
   (* parse the format string *)
   #tDT_TO_STRF := #FMT;
   #pos := FIND(IN1:=#tDT_TO_STRF, IN2:='#');
   WHILE #pos > 0 DO
       (* retrieve format identifier *)
       #f := BYTE_TO_INT("CODE"(STR:=#tDT_TO_STRF, POS:=#pos + 1));
       (* generate the return string according to the format character *)
       #fs := '';
       CASE #f OF
           65 : (* letter A retunrs the year in 4 digits *)
               #fs := DELETE(IN:=S_CONV("YEAR_OF_DATE"(#dx)),L:=1,P:=1);
           66 : (* letter B returns the year in exactly 2 digits *)
               #fs := RIGHT(IN:=DELETE(IN:=S_CONV("YEAR_OF_DATE"(#dx)),L:=1,P:=1),L:=2);
           67 : (* letter C returns the month with 1 or 2 digits *)
               #fs := DELETE(IN:=S_CONV("MONTH_OF_DATE"(#dx)),L:=1,P:=1);
           68 : (* letter D returns the month with exactly 2 digits *)
               #fs := DELETE(IN:=S_CONV("MONTH_OF_DATE"(#dx)),L:=1,P:=1);
               IF LEN(#fs) < 2 THEN #fs := CONCAT(IN1:='0',IN2:=#fs); END_IF;
           69 : (* letter E returns the month with 3 characters *)
               #fs := "MONTH_TO_STRING"(MTH:="MONTH_OF_DATE"(#dx), LANG:=#ly, LX:=3);
           70 : (* letter F returns the month with all characters *)
               #fs := "MONTH_TO_STRING"(MTH:="MONTH_OF_DATE"(#dx), LANG:=#ly, LX:=0);
           71 : (* letter G returns the day with up to 2 digits *)
               #fs := DELETE(IN:=S_CONV("DAY_OF_MONTH"(#dx)),L:=1,P:=1);
           72 : (* letter H returns the day of the month with exactly 2 digits *)
               #fs := DELETE(IN:=S_CONV("DAY_OF_MONTH"(#dx)),L:=1,P:=1);
               IF LEN(#fs) < 2 THEN #fs := CONCAT(IN1:="FILL_FC235", IN2:=#fs); END_IF;
           73 : (* letter I returns the weekday as the number 1..7 1 = monday *)
               #fs := DELETE(IN:=S_CONV("DAY_OF_WEEK"(#dx)),L:=1,P:=1);
           74 : (* letter J returns the weekday in 2 character writing *)
               #fs := "WEEKDAY_TO_STRING"(WDAY:="DAY_OF_WEEK"(#dx), LANG:=#ly, LX:=2);
           75 : (* letter K returns the weekday with all characters *)
               #fs := "WEEKDAY_TO_STRING"(WDAY:="DAY_OF_WEEK"(#dx), LANG:=#ly, LX:=0);
           76 : (* letter L returns AM or PM for the given DateTime *)
               IF #td >= TOD#12:00:00 THEN #fs := 'PM'; ELSE #fs := 'AM'; END_IF;
           77 : (* letter M returns the hour in 1 or 2 digit form 0..24h *)
               #fs := DELETE(IN:=S_CONV("HOUR"(#td)),L:=1,P:=1);
           78 : (* letter N returns the hour in exactly 2 digit form 0..24h *)
               #fs := DELETE(IN:=S_CONV("HOUR"(#td)),L:=1,P:=1);
               IF LEN(#fs) < 2 THEN #fs := CONCAT(IN1:="FILL_FC235", IN2:=#fs); END_IF;
           79 : (* letter O returns the hour in 1 or 2 digit form 0..12h *)
               #tmp := "HOUR"(#td) MOD 12;
               IF #tmp = 0 THEN #tmp := 12; END_IF;
               #fs := DELETE(IN:=S_CONV(#tmp),L:=1,P:=1);
           80 : (* letter P returns the hour in exactly 2 digit form 0..12h *)
               #tmp := "HOUR"(#td) MOD 12;
               IF #tmp = 0 THEN #tmp := 12; END_IF;
               #fs := DELETE(IN:=S_CONV(#tmp),L:=1,P:=1);
               IF LEN(#fs) < 2 THEN #fs := CONCAT(IN1:="FILL_FC235", IN2:=#fs); END_IF;
           81 : (* letter Q returns the minute of the hour in 1 or two digit form *)
               #fs := DELETE(IN:=S_CONV("MINUTE"(#td)),L:=1,P:=1);
           82 : (* letter R returns the minute of the hour in exactly two digit form *)
               #fs := DELETE(IN:=S_CONV("MINUTE"(#td)),L:=1,P:=1);
               IF LEN(#fs) < 2 THEN #fs := CONCAT(IN1:="FILL_FC235", IN2:=#fs); END_IF;
           83 : (* letter S returns the second of the minute in 1 or two digit form *)
               #fs := DELETE(IN:=S_CONV(REAL_TO_INT("SECOND"(#td))),L:=1,P:=1);
           84 : (* letter T returns the second of the minute in exactly two digit form *)
               #fs := DELETE(IN:=S_CONV(REAL_TO_INT("SECOND"(#td))),L:=1,P:=1);
               IF LEN(#fs) < 2 THEN #fs := CONCAT(IN1:="FILL_FC235", IN2:=#fs); END_IF;
           85 : (* letter U returns the milliseconds in 1 to 3 digits *)
               #fs := DELETE(IN:=S_CONV(#MS),L:=1,P:=1);
           86 : (* letter V returns the milliseconds in exactly 3 digit form *)
               #fs := DELETE(IN:=S_CONV(#MS),L:=1,P:=1);
               #fs := CONCAT(IN1:='00',IN2:=#fs);
               #fs := RIGHT(IN:=#fs, L:=3);
           87 : (* letter W returns the day of the month with exactly 2 digits first digit is filled with blank if necessary *)
               #fs := DELETE(IN:=S_CONV("DAY_OF_MONTH"(#dx)),L:=1,P:=1);
               IF LEN(#fs) < 2 THEN #fs := CONCAT(IN1:="BLANK", IN2:=#fs); END_IF;
           88 : (* letter X returns the month with exactly 2 digits first digit is filled with blank if necessary *)
               #fs := DELETE(IN:=S_CONV("MONTH_OF_DATE"(#dx)),L:=1,P:=1);
               IF LEN(#fs) < 2 THEN #fs := CONCAT(IN1:="BLANK", IN2:=#fs); END_IF;
           END_CASE;
       #tDT_TO_STRF := REPLACE(IN1:=#tDT_TO_STRF, IN2:=#fs, L:=2, P:=#pos);
       #pos := FIND(IN1:=#tDT_TO_STRF, IN2:='#');
   END_WHILE;

   #DT_TO_STRF := #tDT_TO_STRF;

   (* revision history
   hm  7. oct. 2008    rev 1.0
       original version

   hm  19. oct. 2008   rev 1.1
       changed language setup constants
   *)
END_FUNCTION

FUNCTION "DWORD_TO_STRB" : String[254]   // FC236, SCL
TITLE = DWORD_TO_STRB
{ S7_Optimized_Access := 'FALSE' }
AUTHOR : hugo
FAMILY : STRINGS
NAME : DW2STRB
VERSION : 1.3
// DWORD_TO_STRINGB converts a DWORD to a String of Bits represented by '0' and '1' s.
// The lowest order bit will be on the right and the high order bit on the left.
   VAR_INPUT
      IN : DWord;
   END_VAR
   VAR_TEMP
      pt : Int;   // pt : POINTER TO BYTE;
      i : Int;
      str : String[32];
      _str AT str : Struct
         length : Byte;
         act_length : Byte;
         str : Array[1..32] of Byte;
      END_STRUCT;
      tIN : DWord;
      _IN AT tIN : Array[0..31] of Bool;
   END_VAR
BEGIN


   #str := #DWORD_TO_STRB;
   #tIN := #IN;

   (* pointer für die ausgabe ermitteln *)
   #pt := 1;    //ADR(DWORD_TO_STRB);
   (* die 8 ausgabecharacter ermitteln und schreiben *)
   FOR #i := 1 TO 32 DO
       #_str.str[#pt] := INT_TO_BYTE(BYTE_TO_INT(BOOL_TO_BYTE(#_IN[7])) + 48);
       #tIN := SHL(IN:=#tIN,N:=1);
       #pt := #pt + 1;
   END_FOR;

   (* der ausgabestring muss nochg mit 32 abgeschlossen werden *)
   #_str.act_length := 32;
   #DWORD_TO_STRB := #str;

   (* revision history
   hm      9.6.2007    rev 1.0     
       original version

   hm      15.dec 2007 rev 1.1
       changed code for better performance

   hm  29. mar. 2008   rev 1.2
       changed STRING to STRING(32)

   hm  20. jun. 2008   rev 1.3
       performance improvement

   *)
END_FUNCTION

FUNCTION "DWORD_TO_STRF" : String[254]   // FC237, SCL
TITLE = DWORD_TO_STRF
{ S7_Optimized_Access := 'FALSE' }
AUTHOR : hugo
FAMILY : STRINGS
NAME : DW2STRF
VERSION : 1.1
// dword_to_strF converts a DWORD, BYTE or Word to a fixed length String.
// the string will be filled with leading zeroes to achieve the fixed length, or if too long, the lowest digits will be used.
// the maximum allowed length is 20 mdigits.
//  
// for example:    dword_to_strf(123,4) = '0123' 
//                 dword_to_strf(123,2) = '23'
// 
// uses: CONCAT [FC2]
//       DI_STRNG [FC5]
//       MID [FC26]
//       LEN [FC21]
   VAR_INPUT
      IN : DWord;
      N : Int;
   END_VAR
   VAR_TEMP
      L : Int;
      temp : String[10];
      temp2 : String[10];
   END_VAR
BEGIN


   (* convert dword to string first and cut to length N *)
   #temp := '0';
   #temp2 := '0';
   #temp := MID(IN:=S_CONV(DWORD_TO_DINT(#IN)), L:=#N, P:=2);
   #L := LEN(#temp);

   WHILE #L < #N DO
       #temp2 := CONCAT(IN1:='0',IN2:=#temp);
       #temp BLKMOV #temp2;
       #L := #L + 1;
   END_WHILE;
   #DWORD_TO_STRF := #temp;


   (* limit N to max 20 characters *)
   //tN := LIMIT(IN1:=0,IN2:=tN,IN3:=20);
   (* convert dword to string first and cut to length N *)
   //str := FIX(DWORD_TO_STRING(in),tN,48,1);

   (* revision history
   hm  26. jan.2007    rev 1.0     
       original version

   hm  29. mar. 2008   rev 1.1
       changed STRING to STRING(20)
       limit the output string to max 20 digits
   *)
END_FUNCTION

FUNCTION "DWORD_TO_STRH" : String[254]   // FC238, SCL
TITLE = DWORD_TO_STRH
{ S7_Optimized_Access := 'FALSE' }
AUTHOR : hugo
FAMILY : STRINGS
NAME : DW2STRH
VERSION : 1.3
// DWORD_TO_STRINGH converts a DWORD to a String of Hexadecimal represented by '0' .. '9' and 'A' .. 'F'.
// The lowest order Character will be on the right and the high order Character on the left.
   VAR_INPUT
      IN : DWord;
   END_VAR
   VAR_TEMP
      i : Int;
      temp : Byte;
      pt : Int;   // pt : POINTER TO BYTE;
      str : String[8];
      _str AT str : Struct
         length : Byte;
         act_length : Byte;
         str : Array[1..8] of Byte;
      END_STRUCT;
      tIN : DWord;
   END_VAR
BEGIN


   #str := #DWORD_TO_STRH;
   #tIN := #IN;

   (* read output adress to pointer *)
   #pt := 8;    //ADR(DWORD_TO_STRH) + 8;
   (* wirte the closing byte for the string *)
   //_str.str[pt]:= 0;

   (* write the 8 hex characters backwards *)
   FOR #i := 1 TO 8 DO;
       (* read the lowest order hex value *)
       #temp := DWORD_TO_BYTE(#tIN AND 16#0000000F);
       (* convert value to hex character *)
       IF BYTE_TO_INT(#temp) <= 9 THEN #temp := INT_TO_BYTE(BYTE_TO_INT(#temp) + 48); ELSE #temp := INT_TO_BYTE(BYTE_TO_INT(#temp) + 55); END_IF;
       (* write character to output string *)
       #_str.str[#pt] := #temp;
       (* shift in for nect hex character *)
       #tIN := SHR(IN:=#tIN,N:=4);
       (* decrement the pointer *)
       #pt := #pt - 1;
   END_FOR;

   #_str.act_length := 8;
   #DWORD_TO_STRH := #str;

   (* code beofre rev 1.2
   FOR i := 1 TO 8 DO
       X := DWORD_TO_BYTE(in AND 2#1111);
       IF X <= 9 THEN X := X + 48; ELSE X := X + 55; END_IF;
       Cx := CHR(X);
       temp := CONCAT(Cx, temp);
       in := SHR(in,4);
   END_FOR;
   DWORD_TO_STRH := temp;
   *)


   (* revision history
   hm  9. jun. 2007    rev 1.0     
       original version 

   hm  11. sep. 2007   rev 1.1
       changed coding for compatibility with twincat, concat cannot support a function as an argument.

   hm  15. dec. 2007    rev 1.2
       changed code for better performance

   hm  29. mar. 2008   rev 1.3
       changed STRING to STRING(8)

   *)
END_FUNCTION

FUNCTION "EXEC" : String[254]   // FC239, SCL
TITLE = EXEC
{ S7_Optimized_Access := 'FALSE' }
AUTHOR : hugo
FAMILY : STRINGS
NAME : EXEC
VERSION : 1.4
// exec executes a mathematical term and returns the result as a string
// the term can only be a simple term without brackets and only one operator
// allowed operastors are: (+, -, *, /, ^, sqrt, sin, cos, tan).
// 
// uses: SETUP [DB1]
//       TEMP [DB7]
//       EQ_STRNG [FC10]
//       R_STRNG [FC30]
//       STRNG_R [FC39]
//       CONCAT [FC2]
//       UPPERCASE [FC288]
//       TO_UPPER [FC284] 
//       TRIM [FC285]
//       FIND [FC11] 
//       REPLACE [FC31] 
//       FINDB_NONUM [FC246]
//       LEFT [FC20]
//       RIGHT [FC32]
//       LEN [FC21]
//       FINDB_NUM [FC247]
   VAR_INPUT
      str : String[254];
   END_VAR
   VAR_TEMP
      pos : Int;
      R1 : Real;
      R2 : Real;
      operator : String[10];
   END_VAR
BEGIN


   "TEMP".STR1 := #str;

   (* extract both numbers and operator *)
   "TEMP".STR2 := "UPPERCASE"("TRIM"("TEMP".STR1));

   #pos := "FINDB_NONUM"("TEMP".STR2);
   IF #pos > 1 THEN #R1 := S_CONV(LEFT(IN:="TEMP".STR2,L:=#pos-1)); END_IF;
   #R2 := S_CONV(RIGHT(IN:="TEMP".STR2,L:=LEN("TEMP".STR2)-#pos));
   "TEMP".STR2 := LEFT(IN:="TEMP".STR2,L:=#pos);
   #pos := "FINDB_NUM"("TEMP".STR2);
   #operator := RIGHT(IN:="TEMP".STR2,L:=LEN("TEMP".STR2) - #pos);
   IF #operator = '' AND LEN("TEMP".STR1) = 0 THEN
       #EXEC := '';
       RETURN;
   ELSIF #operator = '' THEN
       "TEMP".STR2 := "TEMP".STR1;
       RETURN;
   END_IF;
   IF #operator = '^' THEN
       "TEMP".STR2 := S_CONV((#R1**#R2));
   ELSIF #operator = 'SQRT' THEN
       "TEMP".STR2 := S_CONV(SQRT(#R2));
   ELSIF #operator = 'SIN' THEN
       "TEMP".STR2 := S_CONV(SIN(#R2));
   ELSIF #operator = 'COS' THEN
       "TEMP".STR2 := S_CONV(COS(#R2));
   ELSIF #operator = 'TAN' THEN
       "TEMP".STR2 := S_CONV(TAN(#R2));
   ELSIF #operator = '*' THEN
       "TEMP".STR2 := S_CONV(#R1 * #R2);
   ELSIF #operator = '/' THEN
       IF #R2 <> 0 THEN "TEMP".STR2 := S_CONV(#R1 / #R2); ELSE "TEMP".STR2 := 'ERROR'; END_IF;
   ELSIF #operator = '+' THEN
       "TEMP".STR2 := S_CONV(#R1 + #R2);
   ELSIF #operator = '-' THEN
       "TEMP".STR2 := S_CONV(#R1 - #R2);
   ELSE
       "TEMP".STR2 := 'ERROR';
   END_IF;

   IF "TEMP".STR2 = 'ERROR' THEN
       RETURN;
   (* some systems deliver integer instead of real *)
   ELSIF FIND(IN1:="TEMP".STR2,IN2:='.') = 0 THEN
       "TEMP".STR2 := CONCAT(IN1:="TEMP".STR2,IN2:='.0');
   (* some systems deliver n. instead of n.0 ! *)
   ELSIF RIGHT(IN:="TEMP".STR2,L:=1) = '.' THEN
       "TEMP".STR2 := CONCAT(IN1:="TEMP".STR2,IN2:='0');
   END_IF;

   #EXEC := "TEMP".STR2;

   (* revision history

   hm  6.feb 2007      rev 1.1
       cos has to be written in uppercase
       divide by 0 will return an error

   hm  5. mar. 2008    rev 1.2
       add a 0 to the string if a '.' is at the end of the string

   hm  20. mar. 2008   rev 1.3
       make sure the function always returns a real value in the form of x.y

   hm  29. mar. 2008   rev 1.4
       changed STRING to STRING(STRING_LENGTH)
   *)
END_FUNCTION

FUNCTION "FILL" : String[254]   // FC240, SCL
TITLE = FILL
{ S7_Optimized_Access := 'FALSE' }
AUTHOR : hugo
FAMILY : STRINGS
NAME : FILL
VERSION : 1.1
// the function fill creates a string at length L of characters C.
//  
// uses: CONSTANTS [DB6]
//       CONCAT [FC2]
//       CHR_TO_STRING [FC227]
   VAR_INPUT
      C : Byte;
      L : Int;
   END_VAR
   VAR_TEMP
      tFILL : String[254];
      tL : Word;
      _L AT tL : Array[0..15] of Bool;
      i : Int;
      sx : String[1];
   END_VAR
BEGIN


   #sx := "CHR_TO_STRING"(#C);
   (* limit L to maximum 80 characters the length of a standard string *)
   #tL := INT_TO_WORD(LIMIT(MN:=0,IN:=#L,MX:="CONSTANTS".STRING_LENGTH));
   (* create a string of characters to be connected to str *)
   FOR #i := 1 TO 8 DO
       #tFILL := CONCAT(IN1:=#tFILL,IN2:=#tFILL);
       IF #_L[15] THEN #tFILL := CONCAT(IN1:=#tFILL,IN2:=#sx); END_IF;
       #tL := SHL(IN:=#tL,N:=1);
   END_FOR;

   #FILL := #tFILL;


   (* revision histroy
   hm  29. mar. 2008   rev 1.0
       original release

   hm  17. dec. 2008   rev 1.1
       changed function chr to chr_to_string

   *)
END_FUNCTION

FUNCTION "FIND_CHAR" : Int   // FC241, SCL
TITLE = FIND_CHAR
{ S7_Optimized_Access := 'FALSE' }
AUTHOR : hugo
FAMILY : STRINGS
NAME : FCHAR
VERSION : 1.3
// find_char searches str and returns the starting position of the first character that is not a control character.
// control characters are the ascii character 00 .. 31.
// 
// uses: SETUP [DB1]
   VAR_INPUT
      str : String[254];
      _str AT str : Struct
         length : Byte;
         act_length : Byte;
         str : Array[1..254] of Byte;
      END_STRUCT;
      pos : Int;
   END_VAR
   VAR_TEMP
      i : Int;
      stop : Int;
      X : Byte;
   END_VAR
BEGIN


   #stop := BYTE_TO_INT(#_str.act_length);
   FOR #i := MAX(IN1:=#pos,IN2:=1) TO #stop DO
       #X := #_str.str[#i];
       IF BYTE_TO_INT(#X) > 31 AND (("SETUP".EXTENDED_ASCII AND BYTE_TO_INT(#X) <> 127) OR (NOT "SETUP".EXTENDED_ASCII AND BYTE_TO_INT(#X) < 127)) THEN
           #FIND_CHAR := #i;
           RETURN;
       END_IF;
   END_FOR;
   #FIND_CHAR := 0;


   (* revision history
   hm  29. feb 2008    rev 1.0
       original version

   hm  26. mar. 2008   rev 1.1
       char will now accept extended ascii

   hm  29. mar. 2008   rev 1.2
       changed STRING to STRING(STRING_LENGTH)

   hm  21. oct. 2008 rev 1.3
       changes setup constants
       optimized code
   *)
END_FUNCTION

FUNCTION "FIND_CTRL" : Int   // FC242, SCL
TITLE = FIND_CTRL
{ S7_Optimized_Access := 'FALSE' }
AUTHOR : hugo
FAMILY : STRINGS
NAME : FCTRL
VERSION : 1.2
// find_ctrl searches str and returns the starting position of a control character
// control characters are the ascii character 00 .. 31.
   VAR_INPUT
      str : String[254];
      _str AT str : Struct
         length : Byte;
         act_length : Byte;
         str : Array[1..254] of Byte;
      END_STRUCT;
      pos : Int;
   END_VAR
   VAR_TEMP
      i : Int;
      stop : Int;
      x : Byte;
   END_VAR
BEGIN


   #stop := BYTE_TO_INT(#_str.act_length);
   FOR #i := MAX(IN1:=#pos,IN2:=1) TO #stop DO;
       #x := #_str.str[#i];
       IF BYTE_TO_INT(#x) < 32 OR BYTE_TO_INT(#x) = 127 THEN
           #FIND_CTRL := #i;
           RETURN;
       END_IF;
   END_FOR;
   #FIND_CTRL := 0;


   (* revision history
   hm  29. feb 2008    rev 1.0
       original version

   hm  26. mar. 2008   rev 1.1
       character 127 is now recognized as control

   hm  29. mar. 2008   rev 1.2
       changed STRING to STRING(STRING_LENGTH)
   *)
END_FUNCTION

FUNCTION "FIND_NONUM" : Int   // FC243, SCL
TITLE = FIND_NONUM
{ S7_Optimized_Access := 'FALSE' }
AUTHOR : hugo
FAMILY : STRINGS
NAME : FINDNONR
VERSION : 1.3
// find_noNum searches str AND returns the first position which is NOT a number.
// a number is characterized by a letter "0..9" or "."
   VAR_INPUT
      str : String[254];
      _str AT str : Struct
         length : Byte;
         act_length : Byte;
         str : Array[1..254] of Byte;
      END_STRUCT;
      pos : Int;
   END_VAR
   VAR_TEMP
      i : Int;
      end : Int;
      X : Byte;
   END_VAR
BEGIN


   #end := BYTE_TO_INT(#_str.act_length);    //LEN(str);
   FOR #i := MAX(IN1:=#pos,IN2:=1) TO #end DO
       #X := #_str.str[#i];
       IF (BYTE_TO_INT(#X) < 48 AND BYTE_TO_INT(#X) <> 46) OR BYTE_TO_INT(#X) > 57 THEN
           #FIND_NONUM := #i;
           RETURN;
       END_IF;
   END_FOR;
   #FIND_NONUM := 0;


   (* revision history
   hm  6. oct. 2006    rev 1.0
       original version

   hm  29. feb 2008    rev 1.1
       added input pos to start search at position

   hm  29. mar. 2008   rev 1.2
       changed STRING to STRING(STRING_LENGTH)

   hm  21. oct. 2008   rev 1.3
       optimized code

   *)
END_FUNCTION

FUNCTION "FIND_NUM" : Int   // FC244, SCL
TITLE = FIND_NUM
{ S7_Optimized_Access := 'FALSE' }
AUTHOR : hugo
FAMILY : STRINGS
NAME : FINDNR
VERSION : 1.2
// find_Num searches str and returns the starting position of a number
// a number is characterized by a letter "0..9" or "."
   VAR_INPUT
      str : String[254];
      _str AT str : Struct
         length : Byte;
         act_length : Byte;
         str : Array[1..254] of Byte;
      END_STRUCT;
      pos : Int;
   END_VAR
   VAR_TEMP
      i : Int;
      stop : Int;
      X : Byte;
   END_VAR
BEGIN


   #stop := BYTE_TO_INT(#_str.act_length);   //LEN(str);
   FOR #i := MAX(IN1:=#pos,IN2:=1) TO #stop DO;
       #X := #_str.str[#i];
       IF (BYTE_TO_INT(#X) > 47 AND BYTE_TO_INT(#X) < 58) OR BYTE_TO_INT(#X) = 46 THEN
           #FIND_NUM := #i;
           RETURN;
       END_IF;
   END_FOR;
   #FIND_NUM := 0;


   (* revision history
   hm  6. oct. 2006    rev 1.0
       original version

   hm  29. feb 2008    rev 1.1
       added input pos to start search at position

   hm  29. mar. 2008   rev 1.2
       changed STRING to STRING(STRING_LENGTH)

   *)
END_FUNCTION

FUNCTION "FINDB" : Int   // FC245, SCL
TITLE = FINDB
{ S7_Optimized_Access := 'FALSE' }
AUTHOR : hugo
FAMILY : STRINGS
NAME : FINDB
VERSION : 1.3
// the function find searches an str1 for the presence of str2 and returns the first position of str1 of the last presence in instring.
// the function is similar to find except it searches from the right to left.
// a 0 is returned if the string is not found.
//  
// uses: EQ_STRNG [FC10]
//       MID [FC26]
   VAR_INPUT
      str1 : String[254];
      str2 : String[254];
   END_VAR
   VAR_TEMP
      tstr1 : String[254];
      _str1 AT tstr1 : Struct
         length : Byte;
         act_length : Byte;
         str : Array[1..254] of Byte;
      END_STRUCT;
      tstr2 : String[254];
      _str2 AT tstr2 : Struct
         length : Byte;
         act_length : Byte;
         str : Array[1..254] of Byte;
      END_STRUCT;
      pos : Int;
      length : Int;
   END_VAR
BEGIN


   #tstr1 := #str1;
   #tstr2 := #str2;

   #length := BYTE_TO_INT(#_str2.act_length);
   FOR #pos := BYTE_TO_INT(#_str1.act_length) - #length + 1 TO 1 BY -1 DO
       IF MID(IN:=#tstr1,L:=#length,P:=#pos) S_COMP #tstr2 THEN
           #FINDB := #pos;
           RETURN;
       END_IF;
   END_FOR;
   #FINDB := 0;

   (* revision history
   hm  6. oct 2006     rev 1.0
       original version

   hm  15 dec 2007     rev 1.1
       changed code for better performance

   hm  29. feb 2008    rev 1.2
       added findb := 0 for compatibility reasons

   hm  29. mar. 2008   rev 1.3
       changed STRING to STRING(STRING_LENGTH)
   *)
END_FUNCTION

FUNCTION "FINDB_NONUM" : Int   // FC246, SCL
TITLE = FINDB_NONUM
{ S7_Optimized_Access := 'FALSE' }
AUTHOR : hugo
FAMILY : STRINGS
NAME : FINDBNON
VERSION : 1.3
// findB_noNum searches str backwards and returns the last position which is not a number.
// a number is characterized by a letter "0..9" or "."
   VAR_INPUT
      str : String[254];
      _str AT str : Struct
         length : Byte;
         act_length : Byte;
         str : Array[1..254] of Byte;
      END_STRUCT;
   END_VAR
   VAR_TEMP
      pos : Int;
      pt : Int;   // pt : POINTER TO BYTE;
   END_VAR
BEGIN


   #pt := 1 + BYTE_TO_INT(#_str.act_length) - 1;     //ADR(str) + LEN(str) - 1;
   FOR #pos := BYTE_TO_INT(#_str.act_length) TO 1 BY -1 DO;
       IF (BYTE_TO_INT(#_str.str[#pt]) < 48 AND BYTE_TO_INT(#_str.str[#pt]) <> 46) OR BYTE_TO_INT(#_str.str[#pt]) > 57 THEN
           #FINDB_NONUM := #pos;
           RETURN;
       END_IF;
       #pt := #pt - 1;
   END_FOR;
   #FINDB_NONUM := 0;


   (* revision history
   hm  6. oct 2006     rev 1.0
       original version

   hm  29. feb 2008    rev 1.1
       improved performance

   hm  29. mar. 2008   rev 1.2
       changed STRING to STRING(STRING_LENGTH)

   hm  21. oct. 2008   rev 1.3
       optimized code
   *)
END_FUNCTION

FUNCTION "FINDB_NUM" : Int   // FC247, SCL
TITLE = FINDB_NUM
{ S7_Optimized_Access := 'FALSE' }
AUTHOR : hugo
FAMILY : STRINGS
NAME : FINDBNR
VERSION : 1.2
// findB_Num searches str backward and returns the last position of a number
// a number is characterized by a letter "0..9" or "."
   VAR_INPUT
      str : String[254];
      _str AT str : Struct
         length : Byte;
         act_length : Byte;
         str : Array[1..254] of Byte;
      END_STRUCT;
   END_VAR
   VAR_TEMP
      pos : Int;
      pt : Int;   // pt : POINTER TO BYTE;
   END_VAR
BEGIN


   #pt := 1 + BYTE_TO_INT(#_str.act_length) - 1; //ADR(str) + LEN(str) - 1;
   FOR #pos := BYTE_TO_INT(#_str.act_length) TO 1 BY -1 DO;
       IF (BYTE_TO_INT(#_str.str[#pt]) > 47 AND BYTE_TO_INT(#_str.str[#pt]) < 58) OR BYTE_TO_INT(#_str.str[#pt]) = 46 THEN
           #FINDB_NUM := #pos;
           RETURN;
       END_IF;
       #pt := #pt - 1;
   END_FOR;
   #FINDB_NUM := 0;

   (* revision history
   hm  6. oct 2006     rev 1.0
       original version

   hm  29. feb 2008    rev 1.1
       improved performance

   hm  29. mar. 2008   rev 1.2
       changed STRING to STRING(STRING_LENGTH)
   *)
END_FUNCTION

FUNCTION "FINDP" : Int   // FC248, SCL
TITLE = FINDP
{ S7_Optimized_Access := 'FALSE' }
AUTHOR : hugo
FAMILY : STRINGS
NAME : FINDP
VERSION : 1.2
// the function findP searches a string str for the occurence of src beginning at the position pos.
//  
// uses: EQ_STRNG [FC10]
//       MID [FC26]
   VAR_INPUT
      str : String[254];
      src : String[254];
      pos : Int;
   END_VAR
   VAR_TEMP
      tstr : String[254];
      _str AT tstr : Struct
         length : Byte;
         act_length : Byte;
         str : Array[1..254] of Byte;
      END_STRUCT;
      tsrc : String[254];
      _src AT tsrc : Struct
         length : Byte;
         act_length : Byte;
         str : Array[1..254] of Byte;
      END_STRUCT;
      i : Int;
      ls : Int;
      lx : Int;
      stp : Int;
   END_VAR
BEGIN


   #tstr := #str;
   #tsrc := #src;

   #ls := BYTE_TO_INT(#_str.act_length);
   #lx := BYTE_TO_INT(#_src.act_length);
   IF #ls < #lx OR #lx = 0 THEN RETURN; END_IF;
   #stp := #ls - #lx + 1;
   FOR #i := MAX(IN1:=#pos,IN2:=1) TO #stp DO
       IF MID(IN:=#tstr,L:=#lx,P:=#i) = #tsrc THEN
           #FINDP := #i;
           RETURN;
       END_IF;
   END_FOR;
   #FINDP := 0;


   (* revision histroy
   hm  4. feb. 2008    rev 1.0
       original release

   hm  29. feb 2008    rev 1.1
       ADDED MAX(pos,1) in loop initialization

   hm  29. mar. 2008   rev 1.2
       changed STRING to STRING(STRING_LENGTH)
   *)
END_FUNCTION

FUNCTION "FIX" : String[254]   // FC249, SCL
TITLE = FIX
{ S7_Optimized_Access := 'FALSE' }
AUTHOR : hugo
FAMILY : STRINGS
NAME : FIX
VERSION : 1.0
// the function fix truncates a string at length L 
// or if the string is shorter then L it will be filled with ending Spaces till its length = N.
//  
// uses: CONSTANTS [DB6]
//       TEMP [DB7]
//       CONCAT [FC2]
//       LEN [FC21]
//       RIGHT [FC32]
//       LEFT [FC20]
//       FILL [FC240]
//       CHR_TO_STRING [FC227]
   VAR_INPUT
      str : String[254];
      L : Int;
      C : Byte;
      "M" : Int;
   END_VAR
   VAR_TEMP
      N : Int;
      SX : String[254];
   END_VAR
BEGIN


   "TEMP".STR1 := #str;
   "TEMP".STR2 := #FIX;